(* Logix 5000 project; controller MV vendor 1 type 14 code 217 rev 31.11; software revision 31.00; part 4 of 53 *)
(* tags used below, declared in another part *)
   _1s_pulse : BOOL;
   active : BOOL;
   colin : DINT;
   colon_string : STRING;
   hr_string : STRING;
   MC_CH1_CIP_Messages : STRING[20];   // CH1 CIP Scada Messages
   MC_CH1_CIP_Misc : DINT[20];
   MC_CH1_CIP_MiscReal : REAL[20];
   MC_CH1_Delay_For_Data : TIMER;
   MC_CH1_OneShot : BOOL;
   MC_CH1_SaveCIPReport_now : DINT;
   MC_CH1_SaveCIPReport_now_done : DINT;
   MC_CH2_CIP_Messages : STRING[20];   // CH2 CIP Scada Messages
   MC_CH2_CIP_Misc : DINT[20];
   MC_CH2_CIP_MiscReal : REAL[20];
   MC_CH2_Delay_For_Data : TIMER;
   MC_CH2_OneShot : BOOL;
   MC_CH2_SaveCIPReport_now : DINT;
   MC_CH2_SaveCIPReport_now_done : DINT;
   MC_CIP_Default_Messages : STRING[20];
   MC_CIP_temp : INT;
   MC_N100 : INT[255];   // C1_PLC Channel 1 PLC data
   MC_N104 : INT[255];   // CH1 REPORT Channel 1 CIP report file
   MC_N120 : INT[255];   // C2 PLC Channel 2 PLC data
   MC_N124 : INT[255];   // CH2 REPORT Channel 2 CIP report file
   MC_T4 : TIMER[255];   // TIMER
   mn_string : STRING;

        [30].3   // MV 23,Current vessel deferred chilling active
        [16].1   // MV 23,Profile control flag Hold at B.P B
        [16].2   // MV 23,Profile control flag Hold at B.P C
        [16].3   // MV 23,Profile control flag Hold at B.P D
        [16].4   // MV 23,Profile control flag Hold at B.P E
        [0]   // MV 23,FV SYSTEM WORKING BUFFER VESSEL NUMBER
        [21]   // MV 23,Current vessel cold conditioning time
        [2]   // MV 23,TEMPERATURE SETPOINT A. 1/10 DEGREE 'C'
        [30].4   // MV 23,Current vessel final temp.reached
        [16].5   // MV 23,Profile control flag Hold at B.P F
        [16].6   // MV 23,Profile control flag Hold at B.P G
        [4]   // MV 23,TEMPERATURE SETPOINT B. 1/10 DEGREE 'C'
        [6]   // MV 23,TEMPERATURE SETPOINT C. 1/10 DEGREE 'C'
        [8]   // MV 23,TEMPERATURE SETPOINT D. 1/10 DEGREE 'C'
        [27]   // MV 23,CURRENT ELAPSED HOURS *10
        [30].0   // MV 23,Cooling Valve to open
        [24]   // MV 23,Phase 0=off 8=Wait yeast 9=Wait Fill 10=Maturation 11to16=Conditioning
        [10]   // MV 23,TEMPERATURE SETPOINT E. 1/10 DEGREE 'C'
        [12]   // MV 23,TEMPERATURE SETPOINT F. 1/10 DEGREE 'C'
        [14]   // MV 23,TEMPERATURE SETPOINT G. 1/10 DEGREE 'C'
        [15].2   // MV 23,PLC TO FOLLOW RAMP Breakpoints A to B
        [30].6   // MV 23,Current vessel cold cond.temp.reached
        [11]   // MV 23,TEMPERATURE BREAKPOINT F. TIME 1/10 HOURS(ALWAYS=0)
        [13]   // MV 23,TEMPERATURE BREAKPOINT G. TIME 1/10 HOURS(ALWAYS=0)
        [30].5   // MV 23,Current vessel deferred chilling temp.high flag
        [1]   // MV 23,TEMPERATURE BREAKPOINT A. TIME 1/10 HOURS(ALWAYS=0)
        [29].1   // MV 23,Current vessel deferred chilling enabled flag
        [3]   // MV 23,TEMPERATURE BREAKPOINT B. TIME 1/10 HOURS(ALWAYS=0)
        [5]   // MV 23,TEMPERATURE BREAKPOINT C. TIME 1/10 HOURS(ALWAYS=0)
        [7]   // MV 23,TEMPERATURE BREAKPOINT D. TIME 1/10 HOURS(ALWAYS=0)
        [9]   // MV 23,TEMPERATURE BREAKPOINT E. TIME 1/10 HOURS(ALWAYS=0)
        [22]   // MV 23,Current FV total residence time
        [29].0   // MV 23,PC TO SAVE TEMPERATURE DATA
        [15].7   // MV 23,PC>PLC Rousing enabled
        [43]   // MV 23,Current vessel powder type
        [20]   // MV 23,Current FV warm conditioning time
        [15].3   // MV 23,PLC TO USE CONE COOLING JACKET
        [29]   // MV 23,FLAGS - PLC CONTROL
        [25]   // MV 23,ACTUAL TEMPERATURE -DEGREES 'C'*10
        [26]   // MV 23,Calculated Setpoint 1/10 degrees C
        [30].1   // MV 23,Rouser required
        [44]   // MV 23,Current vessel powder amount
        [15]   // MV 23,FLAGS-PROFILE CONTROL
        [28]   // MV 23,CURRENT VOLUME HL*10
   MV_N14 : INT[255] := ([3] := 7);   // ME>PLC Inter PLC comms traf fic outbound
        [3]   // Me>FVSYSTEM Number of cooling valves required by MVSYSTEM
        [2].0   // Me>FVSYSTEM Acknowledgement of request to change MV status to ageing
   MV_N140 : INT[50] := ([0] := 336, [2] := 80, [3] := 1200, [4] := 80, [5] := 2860, [6] := 80, [7] := 5040, [8] := 80, [9] := 6720, [10] := 80, [11] := 8400, [12] := 80, [13] := 32767, [14] := 80, [15] := 148, [17] := -32767, [18] := -32767, [19] := 1680, [20] := 1484, [22] := 3164, [23] := 1, [24] := 10, [25] := 81, [26] := 80, [27] := 1263, [29] := 2, [30] := 24, [32] := 2, [34] := 2, [40] := 2);   // MV 36, CURRENT FV DATA
        [15].4   // MV 36,Profile Control Flags : This is a Maturation Profile
        [15].9   // MV 36,Current vessel deferred chilling manual override
        [15].5   // MV 36,Profile Control Flags : This is a Conditioning Profile
        [36]   // MV 36,Current vessel time to deferred chlling start (hrs.x10)
        [40]   // MV 36,Vessel RoutingStatus 0=Clean,1=Filling,2= Beer,3=Packng1,4=Pac kng2,5=Packng3,6=Ven ting,7=Dirty,8=CIP
        [16].1   // MV 36,Profile control flag Hold at B.P B
        [30].3   // MV 36,Current vessel deferred chilling active
        [16].2   // MV 36,Profile control flag Hold at B.P C
        [16].3   // MV 36,Profile control flag Hold at B.P D
        [16].4   // MV 36,Profile control flag Hold at B.P E
        [16].5   // MV 36,Profile control flag Hold at B.P F
        [16].6   // MV 36,Profile control flag Hold at B.P G
        [0]   // MV 36,FV SYSTEM WORKING BUFFER VESSEL NUMBER
        [21]   // MV 36,Current vessel cold conditioning time
        [2]   // MV 36,TEMPERATURE SETPOINT A. 1/10 DEGREE 'C'
        [30].4   // MV 36,Current vessel final temp.reached
        [4]   // MV 36,TEMPERATURE SETPOINT B. 1/10 DEGREE 'C'
        [6]   // MV 36,TEMPERATURE SETPOINT C. 1/10 DEGREE 'C'
        [8]   // MV 36,TEMPERATURE SETPOINT D. 1/10 DEGREE 'C'
        [27]   // MV 36,CURRENT ELAPSED HOURS *10
        [30].0   // MV 36,Cooling Valve to open
        [10]   // MV 36,TEMPERATURE SETPOINT E. 1/10 DEGREE 'C'
        [12]   // MV 36,TEMPERATURE SETPOINT F. 1/10 DEGREE 'C'
        [14]   // MV 36,TEMPERATURE SETPOINT G. 1/10 DEGREE 'C'
        [24]   // MV 36,Phase 0=off 8=Wait yeast 9=Wait Fill 10=Maturation 11to16=Conditioning
        [15].2   // MV 36,PLC TO FOLLOW RAMP Breakpoints A to B
        [30].6   // MV 36,Current vessel cold cond.temp.reached
        [11]   // MV 36,TEMPERATURE BREAKPOINT F. TIME 1/10 HOURS(ALWAYS=0)
        [13]   // MV 36,TEMPERATURE BREAKPOINT G. TIME 1/10 HOURS(ALWAYS=0)
        [30].5   // MV 36,Current vessel deferred chilling temp.high flag
        [1]   // MV 36,TEMPERATURE BREAKPOINT A. TIME 1/10 HOURS(ALWAYS=0)
        [29].1   // MV 36,Current vessel deferred chilling enabled flag
        [3]   // MV 36,TEMPERATURE BREAKPOINT B. TIME 1/10 HOURS(ALWAYS=0)
        [5]   // MV 36,TEMPERATURE BREAKPOINT C. TIME 1/10 HOURS(ALWAYS=0)
        [7]   // MV 36,TEMPERATURE BREAKPOINT D. TIME 1/10 HOURS(ALWAYS=0)
        [9]   // MV 36,TEMPERATURE BREAKPOINT E. TIME 1/10 HOURS(ALWAYS=0)
        [22]   // MV 36,Current FV total residence time
        [29].0   // MV 36,PC TO SAVE TEMPERATURE DATA
        [15].7   // MV 36,PC>PLC Rousing enabled
        [43]   // MV 36,Current vessel powder type
        [20]   // MV 36,Current FV warm conditioning time
        [29]   // MV 36,FLAGS - PLC CONTROL
        [44]   // MV 36,Current vessel powder amount
        [15].3   // MV 36,PLC TO USE CONE COOLING JACKET
        [30].1   // MV 36,Rouser required
        [25]   // MV 36,ACTUAL TEMPERATURE -DEGREES 'C'*10
        [26]   // MV 36,Calculated Setpoint 1/10 degrees C
        [28]   // MV 36,CURRENT VOLUME HL*10
        [15]   // MV 36,FLAGS-PROFILE CONTROL
   MV_N141 : INT[50] := ([0] := 337, [2] := 100, [3] := 720, [4] := 100, [5] := 1201, [6] := -15, [7] := 4561, [8] := -15, [9] := 6241, [10] := -15, [11] := 6721, [12] := -15, [13] := 32767, [14] := -15, [15] := 164, [17] := -32767, [18] := -32767, [19] := 1680, [20] := 909, [21] := 3968, [22] := 7010, [23] := 1, [24] := 14, [25] := -14, [26] := -15, [27] := 5141, [29] := 2, [30] := 88, [32] := 2, [34] := 2, [40] := 2);   // MV 37, CURRENT FV DATA
        [15].4   // MV 37,Profile Control Flags : This is a Maturation Profile
        [15].9   // MV 37,Current vessel deferred chilling manual override
        [15].5   // MV 37,Profile Control Flags : This is a Conditioning Profile
        [36]   // MV 37,Current vessel time to deferred chlling start (hrs.x10)
        [30].3   // MV 37,Current vessel deferred chilling active
        [40]   // MV 37,Vessel RoutingStatus 0=Clean,1=Filling,2= Beer,3=Packng1,4=Pac kng2,5=Packng3,6=Ven ting,7=Dirty,8=CIP
        [16].1   // MV 37,Profile control flag Hold at B.P B
        [16].2   // MV 37,Profile control flag Hold at B.P C
        [16].3   // MV 37,Profile control flag Hold at B.P D
        [16].4   // MV 37,Profile control flag Hold at B.P E
        [16].5   // MV 37,Profile control flag Hold at B.P F
        [16].6   // MV 37,Profile control flag Hold at B.P G
        [0]   // MV 37,FV SYSTEM WORKING BUFFER VESSEL NUMBER
        [21]   // MV 37,Current vessel cold conditioning time
        [2]   // MV 37,TEMPERATURE SETPOINT A. 1/10 DEGREE 'C'
        [30].4   // MV 37,Current vessel final temp.reached
        [4]   // MV 37,TEMPERATURE SETPOINT B. 1/10 DEGREE 'C'
        [6]   // MV 37,TEMPERATURE SETPOINT C. 1/10 DEGREE 'C'
        [8]   // MV 37,TEMPERATURE SETPOINT D. 1/10 DEGREE 'C'
        [27]   // MV 37,CURRENT ELAPSED HOURS *10
        [30].0   // MV 37,Cooling Valve to open
        [10]   // MV 37,TEMPERATURE SETPOINT E. 1/10 DEGREE 'C'
        [12]   // MV 37,TEMPERATURE SETPOINT F. 1/10 DEGREE 'C'
        [14]   // MV 37,TEMPERATURE SETPOINT G. 1/10 DEGREE 'C'
        [15].2   // MV 37,PLC TO FOLLOW RAMP Breakpoints A to B
        [24]   // MV 37,Phase 0=off 8=Wait yeast 9=Wait Fill 10=Maturation 11to16=Conditioning
        [30].6   // MV 37,Current vessel cold cond.temp.reached
        [11]   // MV 37,TEMPERATURE BREAKPOINT F. TIME 1/10 HOURS(ALWAYS=0)
        [1]   // MV 37,TEMPERATURE BREAKPOINT A. TIME 1/10 HOURS(ALWAYS=0)
        [13]   // MV 37,TEMPERATURE BREAKPOINT G. TIME 1/10 HOURS(ALWAYS=0)
        [30].5   // MV 37,Current vessel deferred chilling temp.high flag
        [29].1   // MV 37,Current vessel deferred chilling enabled flag
        [3]   // MV 37,TEMPERATURE BREAKPOINT B. TIME 1/10 HOURS(ALWAYS=0)
        [5]   // MV 37,TEMPERATURE BREAKPOINT C. TIME 1/10 HOURS(ALWAYS=0)
        [7]   // MV 37,TEMPERATURE BREAKPOINT D. TIME 1/10 HOURS(ALWAYS=0)
        [9]   // MV 37,TEMPERATURE BREAKPOINT E. TIME 1/10 HOURS(ALWAYS=0)
        [22]   // MV 37,Current FV total residence time
        [29].0   // MV 37,PC TO SAVE TEMPERATURE DATA
        [15].7   // MV 37,PC>PLC Rousing enabled
        [43]   // MV 37,Current vessel powder type
        [44]   // MV 37,Current vessel powder amount
        [20]   // MV 37,Current FV warm conditioning time
        [15].3   // MV 37,PLC TO USE CONE COOLING JACKET
        [25]   // MV 37,ACTUAL TEMPERATURE -DEGREES 'C'*10
        [29]   // MV 37,FLAGS - PLC CONTROL
        [26]   // MV 37,Calculated Setpoint 1/10 degrees C
        [30].1   // MV 37,Rouser required
        [15]   // MV 37,FLAGS-PROFILE CONTROL
        [28]   // MV 37,CURRENT VOLUME HL*10
   MV_N142 : INT[50] := ([0] := 338, [2] := 80, [3] := 1200, [4] := 80, [5] := 2860, [6] := 80, [7] := 5040, [8] := 80, [9] := 6720, [10] := 80, [11] := 8400, [12] := 80, [13] := 32767, [14] := 80, [15] := 148, [17] := -32767, [18] := -32767, [19] := 1680, [20] := 1481, [22] := 3161, [23] := 1, [24] := 10, [25] := 81, [26] := 80, [27] := 1275, [29] := 2, [30] := 24, [32] := 2, [34] := 2, [40] := 2);   // MV 38, CURRENT FV DATA
        [15].4   // MV 38,Profile Control Flags : This is a Maturation Profile
        [15].9   // MV 38,Current vessel deferred chilling manual override
        [15].5   // MV 38,Profile Control Flags : This is a Conditioning Profile
        [36]   // MV 38,Current vessel time to deferred chlling start (hrs.x10)
        [30].3   // MV 38,Current vessel deferred chilling active
        [40]   // MV 38,Vessel RoutingStatus 0=Clean,1=Filling,2= Beer,3=Packng1,4=Pac kng2,5=Packng3,6=Ven ting,7=Dirty,8=CIP
        [16].1   // MV 38,Profile control flag Hold at B.P B
        [16].2   // MV 38,Profile control flag Hold at B.P C
        [16].3   // MV 38,Profile control flag Hold at B.P D
        [16].4   // MV 38,Profile control flag Hold at B.P E
        [16].5   // MV 38,Profile control flag Hold at B.P F
        [16].6   // MV 38,Profile control flag Hold at B.P G
        [0]   // MV 38,FV SYSTEM WORKING BUFFER VESSEL NUMBER
        [21]   // MV 38,Current vessel cold conditioning time
        [2]   // MV 38,TEMPERATURE SETPOINT A. 1/10 DEGREE 'C'
        [30].4   // MV 38,Current vessel final temp.reached
        [4]   // MV 38,TEMPERATURE SETPOINT B. 1/10 DEGREE 'C'
        [6]   // MV 38,TEMPERATURE SETPOINT C. 1/10 DEGREE 'C'
        [8]   // MV 38,TEMPERATURE SETPOINT D. 1/10 DEGREE 'C'
        [27]   // MV 38,CURRENT ELAPSED HOURS *10
        [30].0   // MV 38,Cooling Valve to open
        [10]   // MV 38,TEMPERATURE SETPOINT E. 1/10 DEGREE 'C'
        [12]   // MV 38,TEMPERATURE SETPOINT F. 1/10 DEGREE 'C'
        [14]   // MV 38,TEMPERATURE SETPOINT G. 1/10 DEGREE 'C'
        [15].2   // MV 38,PLC TO FOLLOW RAMP Breakpoints A to B
        [30].6   // MV 38,Current vessel cold cond.temp.reached
        [24]   // MV 38,Phase 0=off 8=Wait yeast 9=Wait Fill 10=Maturation 11to16=Conditioning
        [11]   // MV 38,TEMPERATURE BREAKPOINT F. TIME 1/10 HOURS(ALWAYS=0)
        [1]   // MV 38,TEMPERATURE BREAKPOINT A. TIME 1/10 HOURS(ALWAYS=0)
        [13]   // MV 38,TEMPERATURE BREAKPOINT G. TIME 1/10 HOURS(ALWAYS=0)
        [30].5   // MV 38,Current vessel deferred chilling temp.high flag
        [29].1   // MV 38,Current vessel deferred chilling enabled flag
        [3]   // MV 38,TEMPERATURE BREAKPOINT B. TIME 1/10 HOURS(ALWAYS=0)
        [5]   // MV 38,TEMPERATURE BREAKPOINT C. TIME 1/10 HOURS(ALWAYS=0)
        [7]   // MV 38,TEMPERATURE BREAKPOINT D. TIME 1/10 HOURS(ALWAYS=0)
        [9]   // MV 38,TEMPERATURE BREAKPOINT E. TIME 1/10 HOURS(ALWAYS=0)
        [22]   // MV 38,Current FV total residence time
        [29].0   // MV 38,PC TO SAVE TEMPERATURE DATA
        [15].7   // MV 38,PC>PLC Rousing enabled
        [43]   // MV 38,Current vessel powder type
        [44]   // MV 38,Current vessel powder amount
        [15]   // MV 38,FLAGS-PROFILE CONTROL
        [20]   // MV 38,Current FV warm conditioning time
        [15].3   // MV 38,PLC TO USE CONE COOLING JACKET
        [25]   // MV 38,ACTUAL TEMPERATURE -DEGREES 'C'*10
        [29]   // MV 38,FLAGS - PLC CONTROL
        [26]   // MV 38,Calculated Setpoint 1/10 degrees C
        [30].1   // MV 38,Rouser required
        [28]   // MV 38,CURRENT VOLUME HL*10
   MV_N143 : INT[50] := ([0] := 339, [2] := 100, [3] := 720, [4] := 100, [5] := 1201, [6] := -15, [7] := 4561, [8] := -15, [9] := 6241, [10] := -15, [11] := 6721, [12] := -15, [13] := 32767, [14] := -15, [15] := 164, [17] := -32767, [18] := -32767, [19] := 1680, [20] := 720, [21] := 5140, [22] := 7976, [23] := 1, [24] := 15, [25] := -14, [26] := -15, [27] := 6309, [29] := 2, [30] := 88, [32] := 2, [34] := 2, [40] := 2);   // MV 39, CURRENT FV DATA
        [15].4   // MV 39,Profile Control Flags : This is a Maturation Profile
        [15].9   // MV 39,Current vessel deferred chilling manual override
        [15].5   // MV 39,Profile Control Flags : This is a Conditioning Profile
        [36]   // MV 39,Current vessel time to deferred chlling start (hrs.x10)
        [30].3   // MV 39,Current vessel deferred chilling active
        [40]   // MV 39,Vessel RoutingStatus 0=Clean,1=Filling,2= Beer,3=Packng1,4=Pac kng2,5=Packng3,6=Ven ting,7=Dirty,8=CIP
        [16].1   // MV 39,Profile control flag Hold at B.P B
        [16].2   // MV 39,Profile control flag Hold at B.P C
        [16].3   // MV 39,Profile control flag Hold at B.P D
        [16].4   // MV 39,Profile control flag Hold at B.P E
        [16].5   // MV 39,Profile control flag Hold at B.P F
        [16].6   // MV 39,Profile control flag Hold at B.P G
        [0]   // MV 39,FV SYSTEM WORKING BUFFER VESSEL NUMBER
        [21]   // MV 39,Current vessel cold conditioning time
        [2]   // MV 39,TEMPERATURE SETPOINT A. 1/10 DEGREE 'C'
        [30].4   // MV 39,Current vessel final temp.reached
        [4]   // MV 39,TEMPERATURE SETPOINT B. 1/10 DEGREE 'C'
        [6]   // MV 39,TEMPERATURE SETPOINT C. 1/10 DEGREE 'C'
        [8]   // MV 39,TEMPERATURE SETPOINT D. 1/10 DEGREE 'C'
        [27]   // MV 39,CURRENT ELAPSED HOURS *10
        [10]   // MV 39,TEMPERATURE SETPOINT E. 1/10 DEGREE 'C'
        [12]   // MV 39,TEMPERATURE SETPOINT F. 1/10 DEGREE 'C'
        [30].0   // MV 39,Cooling Valve to open
        [14]   // MV 39,TEMPERATURE SETPOINT G. 1/10 DEGREE 'C'
        [15].2   // MV 39,PLC TO FOLLOW RAMP Breakpoints A to B
        [30].6   // MV 39,Current vessel cold cond.temp.reached
        [24]   // MV 39,Phase 0=off 8=Wait yeast 9=Wait Fill 10=Maturation 11to16=Conditioning
        [11]   // MV 39,TEMPERATURE BREAKPOINT F. TIME 1/10 HOURS(ALWAYS=0)
        [1]   // MV 39,TEMPERATURE BREAKPOINT A. TIME 1/10 HOURS(ALWAYS=0)
        [13]   // MV 39,TEMPERATURE BREAKPOINT G. TIME 1/10 HOURS(ALWAYS=0)
        [30].5   // MV 39,Current vessel deferred chilling temp.high flag
        [29].1   // MV 39,Current vessel deferred chilling enabled flag
        [3]   // MV 39,TEMPERATURE BREAKPOINT B. TIME 1/10 HOURS(ALWAYS=0)
        [5]   // MV 39,TEMPERATURE BREAKPOINT C. TIME 1/10 HOURS(ALWAYS=0)
        [7]   // MV 39,TEMPERATURE BREAKPOINT D. TIME 1/10 HOURS(ALWAYS=0)
        [9]   // MV 39,TEMPERATURE BREAKPOINT E. TIME 1/10 HOURS(ALWAYS=0)
        [22]   // MV 39,Current FV total residence time
        [29].0   // MV 39,PC TO SAVE TEMPERATURE DATA
        [15].7   // MV 39,PC>PLC Rousing enabled
        [43]   // MV 39,Current vessel powder type
        [44]   // MV 39,Current vessel powder amount
        [15].3   // MV 39,PLC TO USE CONE COOLING JACKET
        [29]   // MV 39,FLAGS - PLC CONTROL
        [30].1   // MV 39,Rouser required
        [15]   // MV 39,FLAGS-PROFILE CONTROL
        [20]   // MV 39,Current FV warm conditioning time
        [25]   // MV 39,ACTUAL TEMPERATURE -DEGREES 'C'*10
        [26]   // MV 39,Calculated Setpoint 1/10 degrees C
        [28]   // MV 39,CURRENT VOLUME HL*10
   MV_N144 : INT[50] := ([0] := 340, [2] := 80, [3] := 1200, [4] := 80, [5] := 2860, [6] := 80, [7] := 5040, [8] := 80, [9] := 6720, [10] := 80, [11] := 8400, [12] := 80, [13] := 32767, [14] := 80, [15] := 148, [17] := -32767, [18] := -32767, [19] := 1680, [20] := 65, [22] := 1718, [23] := 1, [24] := 10, [25] := 78, [26] := 80, [27] := 65, [30] := 16, [32] := 2, [34] := 2, [36] := 416, [40] := 2);   // MV 40, CURRENT FV DATA
        [15].4   // MV 40,Profile Control Flags : This is a Maturation Profile
        [15].9   // MV 40,Current vessel deferred chilling manual override
        [15].5   // MV 40,Profile Control Flags : This is a Conditioning Profile
        [36]   // MV 40,Current vessel time to deferred chlling start (hrs.x10)
        [30].3   // MV 40,Current vessel deferred chilling active
        [16].1   // MV 40,Profile control flag Hold at B.P B
        [16].2   // MV 40,Profile control flag Hold at B.P C
        [16].3   // MV 40,Profile control flag Hold at B.P D
        [40]   // MV 40,Vessel RoutingStatus 0=Clean,1=Filling,2= Beer,3=Packng1,4=Pac kng2,5=Packng3,6=Ven ting,7=Dirty,8=CIP
        [16].4   // MV 40,Profile control flag Hold at B.P E
        [16].5   // MV 40,Profile control flag Hold at B.P F
        [0]   // MV 40,FV SYSTEM WORKING BUFFER VESSEL NUMBER
        [16].6   // MV 40,Profile control flag Hold at B.P G
        [21]   // MV 40,Current vessel cold conditioning time
        [2]   // MV 40,TEMPERATURE SETPOINT A. 1/10 DEGREE 'C'
        [30].4   // MV 40,Current vessel final temp.reached
        [4]   // MV 40,TEMPERATURE SETPOINT B. 1/10 DEGREE 'C'
        [6]   // MV 40,TEMPERATURE SETPOINT C. 1/10 DEGREE 'C'
        [8]   // MV 40,TEMPERATURE SETPOINT D. 1/10 DEGREE 'C'
        [27]   // MV 40,CURRENT ELAPSED HOURS *10
        [10]   // MV 40,TEMPERATURE SETPOINT E. 1/10 DEGREE 'C'
        [30].0   // MV 40,Cooling Valve to open
        [12]   // MV 40,TEMPERATURE SETPOINT F. 1/10 DEGREE 'C'
        [14]   // MV 40,TEMPERATURE SETPOINT G. 1/10 DEGREE 'C'
        [15].2   // MV 40,PLC TO FOLLOW RAMP Breakpoints A to B
        [30].6   // MV 40,Current vessel cold cond.temp.reached
        [24]   // MV 40,Phase 0=off 8=Wait yeast 9=Wait Fill 10=Maturation 11to16=Conditioning
        [1]   // MV 40,TEMPERATURE BREAKPOINT A. TIME 1/10 HOURS(ALWAYS=0)
        [11]   // MV 40,TEMPERATURE BREAKPOINT F. TIME 1/10 HOURS(ALWAYS=0)
        [29].1   // MV 40,Current vessel deferred chilling enabled flag
        [13]   // MV 40,TEMPERATURE BREAKPOINT G. TIME 1/10 HOURS(ALWAYS=0)
        [30].5   // MV 40,Current vessel deferred chilling temp.high flag
        [3]   // MV 40,TEMPERATURE BREAKPOINT B. TIME 1/10 HOURS(ALWAYS=0)
        [5]   // MV 40,TEMPERATURE BREAKPOINT C. TIME 1/10 HOURS(ALWAYS=0)
        [7]   // MV 40,TEMPERATURE BREAKPOINT D. TIME 1/10 HOURS(ALWAYS=0)
        [9]   // MV 40,TEMPERATURE BREAKPOINT E. TIME 1/10 HOURS(ALWAYS=0)
        [22]   // MV 40,Current FV total residence time
        [29].0   // MV 40,PC TO SAVE TEMPERATURE DATA
        [15].7   // MV 40,PC>PLC Rousing enabled
        [43]   // MV 40,Current vessel powder type
        [44]   // MV 40,Current vessel powder amount
        [15]   // MV 40,FLAGS-PROFILE CONTROL
        [15].3   // MV 40,PLC TO USE CONE COOLING JACKET
        [25]   // MV 40,ACTUAL TEMPERATURE -DEGREES 'C'*10
        [26]   // MV 40,Calculated Setpoint 1/10 degrees C
        [29]   // MV 40,FLAGS - PLC CONTROL
        [30].1   // MV 40,Rouser required
        [20]   // MV 40,Current FV warm conditioning time
        [28]   // MV 40,CURRENT VOLUME HL*10
   MV_N145 : INT[50] := ([0] := 341, [2] := 80, [3] := 1200, [4] := 80, [5] := 2860, [6] := 80, [7] := 5040, [8] := 80, [9] := 6720, [10] := 80, [11] := 8400, [12] := 80, [13] := 32767, [14] := 80, [15] := 148, [17] := -32767, [18] := -32767, [19] := 1680, [20] := 53, [22] := 1716, [23] := 1, [24] := 10, [25] := 78, [26] := 80, [27] := 53, [30] := 16, [32] := 2, [34] := 2, [36] := 428, [40] := 2);   // MV 41, CURRENT FV DATA
        [30].3   // MV 41,Current vessel deferred chilling active
        [15].9   // MV 41,Current vessel deferred chilling manual override
        [15].4   // MV 41,Profile Control Flags : This is a Maturation Profile
        [15].5   // MV 41,Profile Control Flags : This is a Conditioning Profile
        [36]   // MV 41,Current vessel time to deferred chlling start (hrs.x10)
        [16].1   // MV 41,Profile control flag Hold at B.P B
        [16].2   // MV 41,Profile control flag Hold at B.P C
        [16].3   // MV 41,Profile control flag Hold at B.P D
        [16].4   // MV 41,Profile control flag Hold at B.P E
        [16].5   // MV 41,Profile control flag Hold at B.P F
        [16].6   // MV 41,Profile control flag Hold at B.P G
        [40]   // MV 41,Vessel RoutingStatus 0=Clean,1=Filling,2= Beer,3=Packng1,4=Pac kng2,5=Packng3,6=Ven ting,7=Dirty,8=CIP
        [0]   // MV 41,FV SYSTEM WORKING BUFFER VESSEL NUMBER
        [21]   // MV 41,Current vessel cold conditioning time
        [2]   // MV 41,TEMPERATURE SETPOINT A. 1/10 DEGREE 'C'
        [30].4   // MV 41,Current vessel final temp.reached
        [4]   // MV 41,TEMPERATURE SETPOINT B. 1/10 DEGREE 'C'
        [6]   // MV 41,TEMPERATURE SETPOINT C. 1/10 DEGREE 'C'
        [8]   // MV 41,TEMPERATURE SETPOINT D. 1/10 DEGREE 'C'
        [10]   // MV 41,TEMPERATURE SETPOINT E. 1/10 DEGREE 'C'
        [27]   // MV 41,CURRENT ELAPSED HOURS *10
        [30].0   // MV 41,Cooling Valve to open
        [12]   // MV 41,TEMPERATURE SETPOINT F. 1/10 DEGREE 'C'
        [14]   // MV 41,TEMPERATURE SETPOINT G. 1/10 DEGREE 'C'
        [15].2   // MV 41,PLC TO FOLLOW RAMP Breakpoints A to B
        [30].6   // MV 41,Current vessel cold cond.temp.reached
        [24]   // MV 41,Phase 0=off 8=Wait yeast 9=Wait Fill 10=Maturation 11to16=Conditioning
        [11]   // MV 41,TEMPERATURE BREAKPOINT F. TIME 1/10 HOURS(ALWAYS=0)
        [1]   // MV 41,TEMPERATURE BREAKPOINT A. TIME 1/10 HOURS(ALWAYS=0)
        [13]   // MV 41,TEMPERATURE BREAKPOINT G. TIME 1/10 HOURS(ALWAYS=0)
        [29].1   // MV 41,Current vessel deferred chilling enabled flag
        [3]   // MV 41,TEMPERATURE BREAKPOINT B. TIME 1/10 HOURS(ALWAYS=0)
        [30].5   // MV 41,Current vessel deferred chilling temp.high flag
        [5]   // MV 41,TEMPERATURE BREAKPOINT C. TIME 1/10 HOURS(ALWAYS=0)
        [7]   // MV 41,TEMPERATURE BREAKPOINT D. TIME 1/10 HOURS(ALWAYS=0)
        [9]   // MV 41,TEMPERATURE BREAKPOINT E. TIME 1/10 HOURS(ALWAYS=0)
        [22]   // MV 41,Current FV total residence time
        [29].0   // MV 41,PC TO SAVE TEMPERATURE DATA
        [15].7   // MV 41,PC>PLC Rousing enabled
        [43]   // MV 41,Current vessel powder type
        [44]   // MV 41,Current vessel powder amount
        [15]   // MV 41,FLAGS-PROFILE CONTROL
        [15].3   // MV 41,PLC TO USE CONE COOLING JACKET
        [25]   // MV 41,ACTUAL TEMPERATURE -DEGREES 'C'*10
        [26]   // MV 41,Calculated Setpoint 1/10 degrees C
        [29]   // MV 41,FLAGS - PLC CONTROL
        [30].1   // MV 41,Rouser required
        [20]   // MV 41,Current FV warm conditioning time
        [28]   // MV 41,CURRENT VOLUME HL*10
   MV_N146 : INT[50] := ([0] := 342, [1] := -32767, [2] := -32767, [3] := -32767, [4] := -32767, [5] := -32767, [6] := -32767, [7] := -32767, [8] := -32767, [9] := -32767, [10] := -32767, [11] := -32767, [12] := -32767, [13] := -32767, [14] := -32767, [15] := -32767, [16] := -32767, [17] := -32767, [18] := -32767, [19] := -32767, [20] := -32767, [21] := -32767, [22] := -32767, [23] := 2, [25] := 210, [30] := 32, [40] := 7);   // MV 42, CURRENT FV DATA
        [30].3   // MV 42,Current vessel deferred chilling active
        [15].9   // MV 42,Current vessel deferred chilling manual override
        [15].4   // MV 42,Profile Control Flags : This is a Maturation Profile
        [15].5   // MV 42,Profile Control Flags : This is a Conditioning Profile
        [36]   // MV 42,Current vessel time to deferred chlling start (hrs.x10)
        [16].1   // MV 42,Profile control flag Hold at B.P B
        [16].2   // MV 42,Profile control flag Hold at B.P C
        [16].3   // MV 42,Profile control flag Hold at B.P D
        [16].4   // MV 42,Profile control flag Hold at B.P E
        [16].5   // MV 42,Profile control flag Hold at B.P F
        [16].6   // MV 42,Profile control flag Hold at B.P G
        [40]   // MV 42,Vessel RoutingStatus 0=Clean,1=Filling,2= Beer,3=Packng1,4=Pac kng2,5=Packng3,6=Ven ting,7=Dirty,8=CIP
        [0]   // MV 42,FV SYSTEM WORKING BUFFER VESSEL NUMBER
        [21]   // MV 42,Current vessel cold conditioning time
        [2]   // MV 42,TEMPERATURE SETPOINT A. 1/10 DEGREE 'C'
        [30].4   // MV 42,Current vessel final temp.reached
        [4]   // MV 42,TEMPERATURE SETPOINT B. 1/10 DEGREE 'C'
        [6]   // MV 42,TEMPERATURE SETPOINT C. 1/10 DEGREE 'C'
        [8]   // MV 42,TEMPERATURE SETPOINT D. 1/10 DEGREE 'C'
        [10]   // MV 42,TEMPERATURE SETPOINT E. 1/10 DEGREE 'C'
        [12]   // MV 42,TEMPERATURE SETPOINT F. 1/10 DEGREE 'C'
        [14]   // MV 42,TEMPERATURE SETPOINT G. 1/10 DEGREE 'C'
        [27]   // MV 42,CURRENT ELAPSED HOURS *10
        [30].0   // MV 42,Cooling Valve to open
        [15].2   // MV 42,PLC TO FOLLOW RAMP Breakpoints A to B
        [30].6   // MV 42,Current vessel cold cond.temp.reached
        [24]   // MV 42,Phase 0=off 8=Wait yeast 9=Wait Fill 10=Maturation 11to16=Conditioning
        [11]   // MV 42,TEMPERATURE BREAKPOINT F. TIME 1/10 HOURS(ALWAYS=0)
        [13]   // MV 42,TEMPERATURE BREAKPOINT G. TIME 1/10 HOURS(ALWAYS=0)
        [30].5   // MV 42,Current vessel deferred chilling temp.high flag
        [1]   // MV 42,TEMPERATURE BREAKPOINT A. TIME 1/10 HOURS(ALWAYS=0)
        [29].1   // MV 42,Current vessel deferred chilling enabled flag
        [3]   // MV 42,TEMPERATURE BREAKPOINT B. TIME 1/10 HOURS(ALWAYS=0)
        [5]   // MV 42,TEMPERATURE BREAKPOINT C. TIME 1/10 HOURS(ALWAYS=0)
        [22]   // MV 42,Current FV total residence time
        [7]   // MV 42,TEMPERATURE BREAKPOINT D. TIME 1/10 HOURS(ALWAYS=0)
        [9]   // MV 42,TEMPERATURE BREAKPOINT E. TIME 1/10 HOURS(ALWAYS=0)
        [29].0   // MV 42,PC TO SAVE TEMPERATURE DATA
        [15].7   // MV 42,PC>PLC Rousing enabled
        [43]   // MV 42,Current vessel powder type
        [44]   // MV 42,Current vessel powder amount
        [15].3   // MV 42,PLC TO USE CONE COOLING JACKET
        [15]   // MV 42,FLAGS-PROFILE CONTROL
        [25]   // MV 42,ACTUAL TEMPERATURE -DEGREES 'C'*10
        [26]   // MV 42,Calculated Setpoint 1/10 degrees C
        [29]   // MV 42,FLAGS - PLC CONTROL
        [30].1   // MV 42,Rouser required
        [20]   // MV 42,Current FV warm conditioning time
        [28]   // MV 42,CURRENT VOLUME HL*10
   MV_N147 : INT[50] := ([0] := 343, [1] := -32767, [2] := -32767, [3] := -32767, [4] := -32767, [5] := -32767, [6] := -32767, [7] := -32767, [8] := -32767, [9] := -32767, [10] := -32767, [11] := -32767, [12] := -32767, [13] := -32767, [14] := -32767, [15] := -32767, [16] := -32767, [17] := -32767, [18] := -32767, [19] := -32767, [20] := -32767, [21] := -32767, [22] := -32767, [23] := 2, [25] := 212, [30] := 32, [40] := 7);   // MV 43, CURRENT FV DATA
        [30].3   // MV 43,Current vessel deferred chilling active
        [15].4   // MV 43,Profile Control Flags : This is a Maturation Profile
        [15].9   // MV 43,Current vessel deferred chilling manual override
        [15].5   // MV 43,Profile Control Flags : This is a Conditioning Profile
        [36]   // MV 43,Current vessel time to deferred chlling start (hrs.x10)
        [16].1   // MV 43,Profile control flag Hold at B.P B
        [16].2   // MV 43,Profile control flag Hold at B.P C
        [16].3   // MV 43,Profile control flag Hold at B.P D
        [16].4   // MV 43,Profile control flag Hold at B.P E
        [16].5   // MV 43,Profile control flag Hold at B.P F
        [16].6   // MV 43,Profile control flag Hold at B.P G
        [0]   // MV 43,FV SYSTEM WORKING BUFFER VESSEL NUMBER
        [21]   // MV 43,Current vessel cold conditioning time
        [2]   // MV 43,TEMPERATURE SETPOINT A. 1/10 DEGREE 'C'
        [30].4   // MV 43,Current vessel final temp.reached
        [40]   // MV 43,Vessel RoutingStatus 0=Clean,1=Filling,2= Beer,3=Packng1,4=Pac kng2,5=Packng3,6=Ven ting,7=Dirty,8=CIP
        [4]   // MV 43,TEMPERATURE SETPOINT B. 1/10 DEGREE 'C'
        [6]   // MV 43,TEMPERATURE SETPOINT C. 1/10 DEGREE 'C'
        [8]   // MV 43,TEMPERATURE SETPOINT D. 1/10 DEGREE 'C'
        [10]   // MV 43,TEMPERATURE SETPOINT E. 1/10 DEGREE 'C'
        [12]   // MV 43,TEMPERATURE SETPOINT F. 1/10 DEGREE 'C'
        [14]   // MV 43,TEMPERATURE SETPOINT G. 1/10 DEGREE 'C'
        [27]   // MV 43,CURRENT ELAPSED HOURS *10
        [30].0   // MV 43,Cooling Valve to open
        [15].2   // MV 43,PLC TO FOLLOW RAMP Breakpoints A to B
        [30].6   // MV 43,Current vessel cold cond.temp.reached
        [24]   // MV 43,Phase 0=off 8=Wait yeast 9=Wait Fill 10=Maturation 11to16=Conditioning
        [11]   // MV 43,TEMPERATURE BREAKPOINT F. TIME 1/10 HOURS(ALWAYS=0)
        [13]   // MV 43,TEMPERATURE BREAKPOINT G. TIME 1/10 HOURS(ALWAYS=0)
        [30].5   // MV 43,Current vessel deferred chilling temp.high flag
        [1]   // MV 43,TEMPERATURE BREAKPOINT A. TIME 1/10 HOURS(ALWAYS=0)
        [29].1   // MV 43,Current vessel deferred chilling enabled flag
        [3]   // MV 43,TEMPERATURE BREAKPOINT B. TIME 1/10 HOURS(ALWAYS=0)
        [5]   // MV 43,TEMPERATURE BREAKPOINT C. TIME 1/10 HOURS(ALWAYS=0)
        [7]   // MV 43,TEMPERATURE BREAKPOINT D. TIME 1/10 HOURS(ALWAYS=0)
        [9]   // MV 43,TEMPERATURE BREAKPOINT E. TIME 1/10 HOURS(ALWAYS=0)
        [22]   // MV 43,Current FV total residence time
        [15].7   // MV 43,PC>PLC Rousing enabled
        [29].0   // MV 43,PC TO SAVE TEMPERATURE DATA
        [43]   // MV 43,Current vessel powder type
        [44]   // MV 43,Current vessel powder amount
        [15].3   // MV 43,PLC TO USE CONE COOLING JACKET
        [25]   // MV 43,ACTUAL TEMPERATURE -DEGREES 'C'*10
        [26]   // MV 43,Calculated Setpoint 1/10 degrees C
        [15]   // MV 43,FLAGS-PROFILE CONTROL
        [29]   // MV 43,FLAGS - PLC CONTROL
        [30].1   // MV 43,Rouser required
        [20]   // MV 43,Current FV warm conditioning time
        [28]   // MV 43,CURRENT VOLUME HL*10
   MV_N148 : INT[50] := ([0] := 344, [2] := 80, [3] := 1200, [4] := 80, [5] := 2860, [6] := 80, [7] := 5040, [8] := 80, [9] := 6720, [10] := 80, [11] := 8400, [12] := 80, [13] := 32767, [14] := 80, [15] := 148, [17] := -32767, [18] := -32767, [19] := 1680, [20] := 1671, [22] := 3341, [23] := 1, [25] := 211, [30] := 32, [32] := 2, [34] := 2, [40] := 7);   // MV 44, CURRENT FV DATA
        [30].3   // MV 44,Current vessel deferred chilling active
        [15].4   // MV 44,Profile Control Flags : This is a Maturation Profile
        [15].9   // MV 44,Current vessel deferred chilling manual override
        [15].5   // MV 44,Profile Control Flags : This is a Conditioning Profile
        [16].1   // MV 44,Profile control flag Hold at B.P B
        [36]   // MV 44,Current vessel time to deferred chlling start (hrs.x10)
        [16].2   // MV 44,Profile control flag Hold at B.P C
        [16].3   // MV 44,Profile control flag Hold at B.P D
        [16].4   // MV 44,Profile control flag Hold at B.P E
        [16].5   // MV 44,Profile control flag Hold at B.P F
        [16].6   // MV 44,Profile control flag Hold at B.P G
        [0]   // MV 44,FV SYSTEM WORKING BUFFER VESSEL NUMBER
        [21]   // MV 44,Current vessel cold conditioning time
        [2]   // MV 44,TEMPERATURE SETPOINT A. 1/10 DEGREE 'C'
        [30].4   // MV 44,Current vessel final temp.reached
        [4]   // MV 44,TEMPERATURE SETPOINT B. 1/10 DEGREE 'C'
        [6]   // MV 44,TEMPERATURE SETPOINT C. 1/10 DEGREE 'C'
        [24]   // MV 44,Phase 0=off 8=Wait yeast 9=Wait Fill 10=Maturation 11to16=Conditioning
        [8]   // MV 44,TEMPERATURE SETPOINT D. 1/10 DEGREE 'C'
        [40]   // MV 44,Vessel RoutingStatus 0=Clean,1=Filling,2= Beer,3=Packng1,4=Pac kng2,5=Packng3,6=Ven ting,7=Dirty,8=CIP
        [10]   // MV 44,TEMPERATURE SETPOINT E. 1/10 DEGREE 'C'
        [12]   // MV 44,TEMPERATURE SETPOINT F. 1/10 DEGREE 'C'
        [14]   // MV 44,TEMPERATURE SETPOINT G. 1/10 DEGREE 'C'
        [27]   // MV 44,CURRENT ELAPSED HOURS *10
        [15].2   // MV 44,PLC TO FOLLOW RAMP Breakpoints A to B
        [30].0   // MV 44,Cooling Valve to open
        [30].6   // MV 44,Current vessel cold cond.temp.reached
        [11]   // MV 44,TEMPERATURE BREAKPOINT F. TIME 1/10 HOURS(ALWAYS=0)
        [13]   // MV 44,TEMPERATURE BREAKPOINT G. TIME 1/10 HOURS(ALWAYS=0)
        [1]   // MV 44,TEMPERATURE BREAKPOINT A. TIME 1/10 HOURS(ALWAYS=0)
        [30].5   // MV 44,Current vessel deferred chilling temp.high flag
        [29].1   // MV 44,Current vessel deferred chilling enabled flag
        [22]   // MV 44,Current FV total residence time
        [3]   // MV 44,TEMPERATURE BREAKPOINT B. TIME 1/10 HOURS(ALWAYS=0)
        [5]   // MV 44,TEMPERATURE BREAKPOINT C. TIME 1/10 HOURS(ALWAYS=0)
        [15].7   // MV 44,PC>PLC Rousing enabled
        [29].0   // MV 44,PC TO SAVE TEMPERATURE DATA
        [7]   // MV 44,TEMPERATURE BREAKPOINT D. TIME 1/10 HOURS(ALWAYS=0)
        [9]   // MV 44,TEMPERATURE BREAKPOINT E. TIME 1/10 HOURS(ALWAYS=0)
        [43]   // MV 44,Current vessel powder type
        [44]   // MV 44,Current vessel powder amount
        [15].3   // MV 44,PLC TO USE CONE COOLING JACKET
        [25]   // MV 44,ACTUAL TEMPERATURE -DEGREES 'C'*10
        [26]   // MV 44,Calculated Setpoint 1/10 degrees C
        [15]   // MV 44,FLAGS-PROFILE CONTROL
        [29]   // MV 44,FLAGS - PLC CONTROL
        [30].1   // MV 44,Rouser required
        [20]   // MV 44,Current FV warm conditioning time
        [28]   // MV 44,CURRENT VOLUME HL*10
   MV_N149 : INT[50] := ([0] := 345, [2] := 80, [3] := 1200, [4] := 80, [5] := 2860, [6] := 80, [7] := 5040, [8] := 80, [9] := 6720, [10] := 80, [11] := 8400, [12] := 80, [13] := 32767, [14] := 80, [15] := 148, [17] := -32767, [18] := -32767, [19] := 1680, [20] := 82, [22] := 1715, [23] := 1, [24] := 10, [25] := 78, [26] := 80, [27] := 82, [30] := 16, [32] := 2, [34] := 2, [36] := 401, [40] := 2);   // MV 45, CURRENT FV DATA
        [15].4   // MV 45,Profile Control Flags : This is a Maturation Profile
        [15].9   // MV 45,Current vessel deferred chilling manual override
        [30].3   // MV 45,Current vessel deferred chilling active
        [36]   // MV 45,Current vessel time to deferred chlling start (hrs.x10)
        [15].5   // MV 45,Profile Control Flags : This is a Conditioning Profile
        [16].1   // MV 45,Profile control flag Hold at B.P B
        [16].2   // MV 45,Profile control flag Hold at B.P C
        [16].3   // MV 45,Profile control flag Hold at B.P D
        [16].4   // MV 45,Profile control flag Hold at B.P E
        [16].5   // MV 45,Profile control flag Hold at B.P F
        [16].6   // MV 45,Profile control flag Hold at B.P G
        [0]   // MV 45,FV SYSTEM WORKING BUFFER VESSEL NUMBER
        [21]   // MV 45,Current vessel cold conditioning time
        [2]   // MV 45,TEMPERATURE SETPOINT A. 1/10 DEGREE 'C'
        [24]   // MV 45,Phase 0=off 8=Wait yeast 9=Wait Fill 10=Maturation 11to16=Conditioning
        [30].4   // MV 45,Current vessel final temp.reached
        [4]   // MV 45,TEMPERATURE SETPOINT B. 1/10 DEGREE 'C'
        [6]   // MV 45,TEMPERATURE SETPOINT C. 1/10 DEGREE 'C'
        [8]   // MV 45,TEMPERATURE SETPOINT D. 1/10 DEGREE 'C'
        [40]   // MV 45,Vessel RoutingStatus 0=Clean,1=Filling,2= Beer,3=Packng1,4=Pac kng2,5=Packng3,6=Ven ting,7=Dirty,8=CIP
        [10]   // MV 45,TEMPERATURE SETPOINT E. 1/10 DEGREE 'C'
        [12]   // MV 45,TEMPERATURE SETPOINT F. 1/10 DEGREE 'C'
        [14]   // MV 45,TEMPERATURE SETPOINT G. 1/10 DEGREE 'C'
        [15].2   // MV 45,PLC TO FOLLOW RAMP Breakpoints A to B
        [30].6   // MV 45,Current vessel cold cond.temp.reached
        [11]   // MV 45,TEMPERATURE BREAKPOINT F. TIME 1/10 HOURS(ALWAYS=0)
        [13]   // MV 45,TEMPERATURE BREAKPOINT G. TIME 1/10 HOURS(ALWAYS=0)
        [27]   // MV 45,CURRENT ELAPSED HOURS *10
        [30].0   // MV 45,Cooling Valve to open
        [30].5   // MV 45,Current vessel deferred chilling temp.high flag
        [1]   // MV 45,TEMPERATURE BREAKPOINT A. TIME 1/10 HOURS(ALWAYS=0)
        [29].1   // MV 45,Current vessel deferred chilling enabled flag
        [3]   // MV 45,TEMPERATURE BREAKPOINT B. TIME 1/10 HOURS(ALWAYS=0)
        [5]   // MV 45,TEMPERATURE BREAKPOINT C. TIME 1/10 HOURS(ALWAYS=0)
        [7]   // MV 45,TEMPERATURE BREAKPOINT D. TIME 1/10 HOURS(ALWAYS=0)
        [9]   // MV 45,TEMPERATURE BREAKPOINT E. TIME 1/10 HOURS(ALWAYS=0)
        [22]   // MV 45,Current FV total residence time
        [15].7   // MV 45,PC>PLC Rousing enabled
        [29].0   // MV 45,PC TO SAVE TEMPERATURE DATA
        [43]   // MV 45,Current vessel powder type
        [44]   // MV 45,Current vessel powder amount
        [15].3   // MV 45,PLC TO USE CONE COOLING JACKET
        [25]   // MV 45,ACTUAL TEMPERATURE -DEGREES 'C'*10
        [15]   // MV 45,FLAGS-PROFILE CONTROL
        [26]   // MV 45,Calculated Setpoint 1/10 degrees C
        [29]   // MV 45,FLAGS - PLC CONTROL
        [30].1   // MV 45,Rouser required
        [20]   // MV 45,Current FV warm conditioning time
        [28]   // MV 45,CURRENT VOLUME HL*10
   MV_N15 : INT[255] := ([0] := 8192, [2] := 16, [3] := 14, [4] := 137, [8] := 23, [14] := 14641, [15] := 11826, [16] := 13873, [17] := 11832, [18] := 12338, [19] := 13102, [20] := 49, [64] := 145);   // COMMS_CTRL Inter PLC comms inte rnal working regs
        [64]   // Pointer to MV data file
        [63].0   // Status change request processing oneshot
   MV_N150 : INT[50] := ([0] := 346, [2] := 80, [3] := 1200, [4] := 80, [5] := 2860, [6] := 80, [7] := 5040, [8] := 80, [9] := 6720, [10] := 80, [11] := 8400, [12] := 80, [13] := 32767, [14] := 80, [15] := 148, [17] := -32767, [18] := -32767, [19] := 1680, [20] := 23726, [22] := 25406, [23] := 3, [25] := 213, [30] := 32, [40] := 7);   // MV 36, CURRENT FV DATA
        [15].9   // MV 36,Current vessel deferred chilling manual override
        [15].4   // MV 36,Profile Control Flags : This is a Maturation Profile
        [24]   // MV 36,Phase 0=off 8=Wait yeast 9=Wait Fill 10=Maturation 11to16=Conditioning
        [30].3   // MV 36,Current vessel deferred chilling active
        [36]   // MV 36,Current vessel time to deferred chlling start (hrs.x10)
        [16].1   // MV 36,Profile control flag Hold at B.P B
        [16].2   // MV 36,Profile control flag Hold at B.P C
        [16].3   // MV 36,Profile control flag Hold at B.P D
        [16].4   // MV 36,Profile control flag Hold at B.P E
        [11]   // MV 36,TEMPERATURE BREAKPOINT F. TIME 1/10 HOURS(ALWAYS=0)
        [15].5   // MV 36,Profile Control Flags : This is a Conditioning Profile
        [16].5   // MV 36,Profile control flag Hold at B.P F
        [16].6   // MV 36,Profile control flag Hold at B.P G
        [0]   // MV 36,FV SYSTEM WORKING BUFFER VESSEL NUMBER
        [21]   // MV 36,Current vessel cold conditioning time
        [2]   // MV 36,TEMPERATURE SETPOINT A. 1/10 DEGREE 'C'
        [30].4   // MV 36,Current vessel final temp.reached
        [4]   // MV 36,TEMPERATURE SETPOINT B. 1/10 DEGREE 'C'
        [6]   // MV 36,TEMPERATURE SETPOINT C. 1/10 DEGREE 'C'
        [8]   // MV 36,TEMPERATURE SETPOINT D. 1/10 DEGREE 'C'
        [40]   // MV 36,Vessel RoutingStatus 0=Clean,1=Filling,2= Beer,3=Packng1,4=Pac kng2,5=Packng3,6=Ven ting,7=Dirty,8=CIP